HMI tags "DB_SDC_ERROR_STAT_EMS011"
   "DB_SDC_ERRORS_STAT_ER_AKT[11].ER_TRIGER" : Word = PLC DB_SDC_ERRORS_STAT.ER_AKT[11].ER_TRIGER AT %DB3724.DBW28680, 1 s
   "DB_SDC_ERRORS_STAT_ER_AKT[11].ER_STAT[1].DRIVE_POS" : DInt = PLC DB_SDC_ERRORS_STAT.ER_AKT[11].ER_STAT[1].DRIVE_POS AT %DB3724.DBD28686, 1 s
   "DB_SDC_ERRORS_STAT_ER_AKT[11].ER_STAT[1].ERROR" : Int = PLC DB_SDC_ERRORS_STAT.ER_AKT[11].ER_STAT[1].ERROR AT %DB3724.DBW28692, 1 s
   "DB_SDC_ERRORS_STAT_ER_AKT[11].ER_STAT[2].DRIVE_POS" : DInt = PLC DB_SDC_ERRORS_STAT.ER_AKT[11].ER_STAT[2].DRIVE_POS AT %DB3724.DBD28702, 1 s
   "DB_SDC_ERRORS_STAT_ER_AKT[11].ER_STAT[2].ERROR" : Int = PLC DB_SDC_ERRORS_STAT.ER_AKT[59].ER_STAT[4].ERROR AT %DB3724.DBW28708, 1 s
   "DB_SDC_ERRORS_STAT_ER_AKT[11].ER_STAT[3].DRIVE_POS" : DInt = PLC DB_SDC_ERRORS_STAT.ER_AKT[11].ER_STAT[3].DRIVE_POS AT %DB3724.DBD28718, 1 s
   "DB_SDC_ERRORS_STAT_ER_AKT[11].ER_STAT[3].ERROR" : Int = PLC DB_SDC_ERRORS_STAT.ER_AKT[11].ER_STAT[3].ERROR AT %DB3724.DBW28724, 1 s
   "DB_SDC_ERRORS_STAT_ER_AKT[11].ER_STAT[4].DRIVE_POS" : DInt = PLC DB_SDC_ERRORS_STAT.ER_AKT[11].ER_STAT[4].DRIVE_POS AT %DB3724.DBD28734, 1 s
   "DB_SDC_ERRORS_STAT_ER_AKT[11].ER_STAT[4].ERROR" : Int = PLC DB_SDC_ERRORS_STAT.ER_AKT[11].ER_STAT[4].ERROR AT %DB3724.DBW28740, 1 s

HMI tags "DB_SDC_ERROR_STAT_EMS012"
   "DB_SDC_ERRORS_STAT_ER_AKT[12].ER_TRIGER" : Word = PLC DB_SDC_ERRORS_STAT.ER_AKT[12].ER_TRIGER AT %DB3724.DBW28746, 1 s
   "DB_SDC_ERRORS_STAT_ER_AKT[12].ER_STAT[1].DRIVE_POS" : DInt = PLC DB_SDC_ERRORS_STAT.ER_AKT[12].ER_STAT[1].DRIVE_POS AT %DB3724.DBD28752, 1 s
   "DB_SDC_ERRORS_STAT_ER_AKT[12].ER_STAT[1].ERROR" : Int = PLC DB_SDC_ERRORS_STAT.ER_AKT[12].ER_STAT[1].ERROR AT %DB3724.DBW28758, 1 s
   "DB_SDC_ERRORS_STAT_ER_AKT[12].ER_STAT[2].DRIVE_POS" : DInt = PLC DB_SDC_ERRORS_STAT.ER_AKT[12].ER_STAT[2].DRIVE_POS AT %DB3724.DBD28768, 1 s
   "DB_SDC_ERRORS_STAT_ER_AKT[12].ER_STAT[2].ERROR" : Int = PLC DB_SDC_ERRORS_STAT.ER_AKT[12].ER_STAT[2].ERROR AT %DB3724.DBW28774, 1 s
   "DB_SDC_ERRORS_STAT_ER_AKT[12].ER_STAT[3].DRIVE_POS" : DInt = PLC DB_SDC_ERRORS_STAT.ER_AKT[12].ER_STAT[3].DRIVE_POS AT %DB3724.DBD28784, 1 s
   "DB_SDC_ERRORS_STAT_ER_AKT[12].ER_STAT[3].ERROR" : Int = PLC DB_SDC_ERRORS_STAT.ER_AKT[12].ER_STAT[3].ERROR AT %DB3724.DBW28790, 1 s
   "DB_SDC_ERRORS_STAT_ER_AKT[12].ER_STAT[4].DRIVE_POS" : DInt = PLC DB_SDC_ERRORS_STAT.ER_AKT[12].ER_STAT[4].DRIVE_POS AT %DB3724.DBD28800, 1 s
   "DB_SDC_ERRORS_STAT_ER_AKT[12].ER_STAT[4].ERROR" : Int = PLC DB_SDC_ERRORS_STAT.ER_AKT[12].ER_STAT[4].ERROR AT %DB3724.DBW28806, 1 s

HMI tags "DB_SDC_ERROR_STAT_EMS013"
   "DB_SDC_ERRORS_STAT_ER_AKT[13].ER_TRIGER" : Word = PLC DB_SDC_ERRORS_STAT.ER_AKT[13].ER_TRIGER AT %DB3724.DBW28812, 1 s
   "DB_SDC_ERRORS_STAT_ER_AKT[13].ER_STAT[1].DRIVE_POS" : DInt = PLC DB_SDC_ERRORS_STAT.ER_AKT[13].ER_STAT[1].DRIVE_POS AT %DB3724.DBD28818, 1 s
   "DB_SDC_ERRORS_STAT_ER_AKT[13].ER_STAT[1].ERROR" : Int = PLC DB_SDC_ERRORS_STAT.ER_AKT[13].ER_STAT[1].ERROR AT %DB3724.DBW28824, 1 s
   "DB_SDC_ERRORS_STAT_ER_AKT[13].ER_STAT[2].DRIVE_POS" : DInt = PLC DB_SDC_ERRORS_STAT.ER_AKT[13].ER_STAT[2].DRIVE_POS AT %DB3724.DBD28834, 1 s
   "DB_SDC_ERRORS_STAT_ER_AKT[13].ER_STAT[2].ERROR" : Int = PLC DB_SDC_ERRORS_STAT.ER_AKT[13].ER_STAT[2].ERROR AT %DB3724.DBW28840, 1 s
   "DB_SDC_ERRORS_STAT_ER_AKT[13].ER_STAT[3].DRIVE_POS" : DInt = PLC DB_SDC_ERRORS_STAT.ER_AKT[13].ER_STAT[3].DRIVE_POS AT %DB3724.DBD28850, 1 s
   "DB_SDC_ERRORS_STAT_ER_AKT[13].ER_STAT[3].ERROR" : Int = PLC DB_SDC_ERRORS_STAT.ER_AKT[13].ER_STAT[3].ERROR AT %DB3724.DBW28856, 1 s
   "DB_SDC_ERRORS_STAT_ER_AKT[13].ER_STAT[4].DRIVE_POS" : DInt = PLC DB_SDC_ERRORS_STAT.ER_AKT[13].ER_STAT[4].DRIVE_POS AT %DB3724.DBD28866, 1 s
   "DB_SDC_ERRORS_STAT_ER_AKT[13].ER_STAT[4].ERROR" : Int = PLC DB_SDC_ERRORS_STAT.ER_AKT[13].ER_STAT[4].ERROR AT %DB3724.DBW28872, 1 s

HMI tags "DB_SDC_ERROR_STAT_EMS014"
   "DB_SDC_ERRORS_STAT_ER_AKT[14].ER_TRIGER" : Word = PLC DB_SDC_ERRORS_STAT.ER_AKT[14].ER_TRIGER AT %DB3724.DBW28878, 1 s
   "DB_SDC_ERRORS_STAT_ER_AKT[14].ER_STAT[1].DRIVE_POS" : DInt = PLC DB_SDC_ERRORS_STAT.ER_AKT[14].ER_STAT[1].DRIVE_POS AT %DB3724.DBD28884, 1 s
   "DB_SDC_ERRORS_STAT_ER_AKT[14].ER_STAT[1].ERROR" : Int = PLC DB_SDC_ERRORS_STAT.ER_AKT[14].ER_STAT[1].ERROR AT %DB3724.DBW28890, 1 s
   "DB_SDC_ERRORS_STAT_ER_AKT[14].ER_STAT[2].DRIVE_POS" : DInt = PLC DB_SDC_ERRORS_STAT.ER_AKT[14].ER_STAT[2].DRIVE_POS AT %DB3724.DBD28900, 1 s
   "DB_SDC_ERRORS_STAT_ER_AKT[14].ER_STAT[2].ERROR" : Int = PLC DB_SDC_ERRORS_STAT.ER_AKT[14].ER_STAT[2].ERROR AT %DB3724.DBW28906, 1 s
   "DB_SDC_ERRORS_STAT_ER_AKT[14].ER_STAT[3].DRIVE_POS" : DInt = PLC DB_SDC_ERRORS_STAT.ER_AKT[14].ER_STAT[3].DRIVE_POS AT %DB3724.DBD28916, 1 s
   "DB_SDC_ERRORS_STAT_ER_AKT[14].ER_STAT[3].ERROR" : Int = PLC DB_SDC_ERRORS_STAT.ER_AKT[14].ER_STAT[3].ERROR AT %DB3724.DBW28922, 1 s
   "DB_SDC_ERRORS_STAT_ER_AKT[14].ER_STAT[4].DRIVE_POS" : DInt = PLC DB_SDC_ERRORS_STAT.ER_AKT[14].ER_STAT[4].DRIVE_POS AT %DB3724.DBD28932, 1 s
   "DB_SDC_ERRORS_STAT_ER_AKT[14].ER_STAT[4].ERROR" : Int = PLC DB_SDC_ERRORS_STAT.ER_AKT[14].ER_STAT[4].ERROR AT %DB3724.DBW28938, 1 s

HMI tags "DB_SDC_ERROR_STAT_EMS015"
   "DB_SDC_ERRORS_STAT_ER_AKT[15].ER_TRIGER" : Word = PLC DB_SDC_ERRORS_STAT.ER_AKT[15].ER_TRIGER AT %DB3724.DBW28944, 1 s
   "DB_SDC_ERRORS_STAT_ER_AKT[15].ER_STAT[1].DRIVE_POS" : DInt = PLC DB_SDC_ERRORS_STAT.ER_AKT[15].ER_STAT[1].DRIVE_POS AT %DB3724.DBD28950, 1 s
   "DB_SDC_ERRORS_STAT_ER_AKT[15].ER_STAT[1].ERROR" : Int = PLC DB_SDC_ERRORS_STAT.ER_AKT[15].ER_STAT[1].ERROR AT %DB3724.DBW28956, 1 s
   "DB_SDC_ERRORS_STAT_ER_AKT[15].ER_STAT[2].DRIVE_POS" : DInt = PLC DB_SDC_ERRORS_STAT.ER_AKT[15].ER_STAT[2].DRIVE_POS AT %DB3724.DBD28966, 1 s
   "DB_SDC_ERRORS_STAT_ER_AKT[15].ER_STAT[2].ERROR" : Int = PLC DB_SDC_ERRORS_STAT.ER_AKT[15].ER_STAT[2].ERROR AT %DB3724.DBW28972, 1 s
   "DB_SDC_ERRORS_STAT_ER_AKT[15].ER_STAT[3].DRIVE_POS" : DInt = PLC DB_SDC_ERRORS_STAT.ER_AKT[15].ER_STAT[3].DRIVE_POS AT %DB3724.DBD28982, 1 s
   "DB_SDC_ERRORS_STAT_ER_AKT[15].ER_STAT[3].ERROR" : Int = PLC DB_SDC_ERRORS_STAT.ER_AKT[15].ER_STAT[3].ERROR AT %DB3724.DBW28988, 1 s
   "DB_SDC_ERRORS_STAT_ER_AKT[15].ER_STAT[4].DRIVE_POS" : DInt = PLC DB_SDC_ERRORS_STAT.ER_AKT[15].ER_STAT[4].DRIVE_POS AT %DB3724.DBD28998, 1 s
   "DB_SDC_ERRORS_STAT_ER_AKT[15].ER_STAT[4].ERROR" : Int = PLC DB_SDC_ERRORS_STAT.ER_AKT[15].ER_STAT[4].ERROR AT %DB3724.DBW29004, 1 s

HMI tags "DB_SDC_ERROR_STAT_EMS016"
   "DB_SDC_ERRORS_STAT_ER_AKT[16].ER_TRIGER" : Word = PLC DB_SDC_ERRORS_STAT.ER_AKT[16].ER_TRIGER AT %DB3724.DBW29010, 1 s
   "DB_SDC_ERRORS_STAT_ER_AKT[16].ER_STAT[1].DRIVE_POS" : DInt = PLC DB_SDC_ERRORS_STAT.ER_AKT[16].ER_STAT[1].DRIVE_POS AT %DB3724.DBD29016, 1 s
   "DB_SDC_ERRORS_STAT_ER_AKT[16].ER_STAT[1].ERROR" : Int = PLC DB_SDC_ERRORS_STAT.ER_AKT[16].ER_STAT[1].ERROR AT %DB3724.DBW29022, 1 s
   "DB_SDC_ERRORS_STAT_ER_AKT[16].ER_STAT[2].DRIVE_POS" : DInt = PLC DB_SDC_ERRORS_STAT.ER_AKT[16].ER_STAT[2].DRIVE_POS AT %DB3724.DBD29032, 1 s
   "DB_SDC_ERRORS_STAT_ER_AKT[16].ER_STAT[2].ERROR" : Int = PLC DB_SDC_ERRORS_STAT.ER_AKT[16].ER_STAT[2].ERROR AT %DB3724.DBW29038, 1 s
   "DB_SDC_ERRORS_STAT_ER_AKT[16].ER_STAT[3].DRIVE_POS" : DInt = PLC DB_SDC_ERRORS_STAT.ER_AKT[16].ER_STAT[3].DRIVE_POS AT %DB3724.DBD29048, 1 s
   "DB_SDC_ERRORS_STAT_ER_AKT[16].ER_STAT[3].ERROR" : Int = PLC DB_SDC_ERRORS_STAT.ER_AKT[16].ER_STAT[3].ERROR AT %DB3724.DBW29054, 1 s
   "DB_SDC_ERRORS_STAT_ER_AKT[16].ER_STAT[4].DRIVE_POS" : DInt = PLC DB_SDC_ERRORS_STAT.ER_AKT[16].ER_STAT[4].DRIVE_POS AT %DB3724.DBD29064, 1 s
   "DB_SDC_ERRORS_STAT_ER_AKT[16].ER_STAT[4].ERROR" : Int = PLC DB_SDC_ERRORS_STAT.ER_AKT[16].ER_STAT[4].ERROR AT %DB3724.DBW29070, 1 s

HMI tags "DB_SDC_ERROR_STAT_EMS017"
   "DB_SDC_ERRORS_STAT_ER_AKT[17].ER_TRIGER" : Word = PLC DB_SDC_ERRORS_STAT.ER_AKT[17].ER_TRIGER AT %DB3724.DBW29076, 1 s
   "DB_SDC_ERRORS_STAT_ER_AKT[17].ER_STAT[1].DRIVE_POS" : DInt = PLC DB_SDC_ERRORS_STAT.ER_AKT[17].ER_STAT[1].DRIVE_POS AT %DB3724.DBD29082, 1 s
   "DB_SDC_ERRORS_STAT_ER_AKT[17].ER_STAT[1].ERROR" : Int = PLC DB_SDC_ERRORS_STAT.ER_AKT[17].ER_STAT[1].ERROR AT %DB3724.DBW29088, 1 s
   "DB_SDC_ERRORS_STAT_ER_AKT[17].ER_STAT[2].DRIVE_POS" : DInt = PLC DB_SDC_ERRORS_STAT.ER_AKT[17].ER_STAT[2].DRIVE_POS AT %DB3724.DBD29098, 1 s
   "DB_SDC_ERRORS_STAT_ER_AKT[17].ER_STAT[2].ERROR" : Int = PLC DB_SDC_ERRORS_STAT.ER_AKT[17].ER_STAT[2].ERROR AT %DB3724.DBW29104, 1 s
   "DB_SDC_ERRORS_STAT_ER_AKT[17].ER_STAT[3].DRIVE_POS" : DInt = PLC DB_SDC_ERRORS_STAT.ER_AKT[17].ER_STAT[3].DRIVE_POS AT %DB3724.DBD29114, 1 s
   "DB_SDC_ERRORS_STAT_ER_AKT[17].ER_STAT[3].ERROR" : Int = PLC DB_SDC_ERRORS_STAT.ER_AKT[17].ER_STAT[3].ERROR AT %DB3724.DBW29120, 1 s
   "DB_SDC_ERRORS_STAT_ER_AKT[17].ER_STAT[4].DRIVE_POS" : DInt = PLC DB_SDC_ERRORS_STAT.ER_AKT[17].ER_STAT[4].DRIVE_POS AT %DB3724.DBD29130, 1 s
   "DB_SDC_ERRORS_STAT_ER_AKT[17].ER_STAT[4].ERROR" : Int = PLC DB_SDC_ERRORS_STAT.ER_AKT[17].ER_STAT[4].ERROR AT %DB3724.DBW29136, 1 s

HMI tags "DB_SDC_ERROR_STAT_EMS018"
   "DB_SDC_ERRORS_STAT_ER_AKT[18].ER_TRIGER" : Word = PLC DB_SDC_ERRORS_STAT.ER_AKT[18].ER_TRIGER AT %DB3724.DBW29142, 1 s
   "DB_SDC_ERRORS_STAT_ER_AKT[18].ER_STAT[1].DRIVE_POS" : DInt = PLC DB_SDC_ERRORS_STAT.ER_AKT[18].ER_STAT[1].DRIVE_POS AT %DB3724.DBD29148, 1 s
   "DB_SDC_ERRORS_STAT_ER_AKT[18].ER_STAT[1].ERROR" : Int = PLC DB_SDC_ERRORS_STAT.ER_AKT[18].ER_STAT[1].ERROR AT %DB3724.DBW29154, 1 s
   "DB_SDC_ERRORS_STAT_ER_AKT[18].ER_STAT[2].DRIVE_POS" : DInt = PLC DB_SDC_ERRORS_STAT.ER_AKT[18].ER_STAT[2].DRIVE_POS AT %DB3724.DBD29164, 1 s
   "DB_SDC_ERRORS_STAT_ER_AKT[18].ER_STAT[2].ERROR" : Int = PLC DB_SDC_ERRORS_STAT.ER_AKT[18].ER_STAT[2].ERROR AT %DB3724.DBW29170, 1 s
   "DB_SDC_ERRORS_STAT_ER_AKT[18].ER_STAT[3].DRIVE_POS" : DInt = PLC DB_SDC_ERRORS_STAT.ER_AKT[18].ER_STAT[3].DRIVE_POS AT %DB3724.DBD29180, 1 s
   "DB_SDC_ERRORS_STAT_ER_AKT[18].ER_STAT[3].ERROR" : Int = PLC DB_SDC_ERRORS_STAT.ER_AKT[18].ER_STAT[3].ERROR AT %DB3724.DBW29186, 1 s
   "DB_SDC_ERRORS_STAT_ER_AKT[18].ER_STAT[4].DRIVE_POS" : DInt = PLC DB_SDC_ERRORS_STAT.ER_AKT[18].ER_STAT[4].DRIVE_POS AT %DB3724.DBD29196, 1 s
   "DB_SDC_ERRORS_STAT_ER_AKT[18].ER_STAT[4].ERROR" : Int = PLC DB_SDC_ERRORS_STAT.ER_AKT[18].ER_STAT[4].ERROR AT %DB3724.DBW29202, 1 s

HMI tags "DB_SDC_ERROR_STAT_EMS019"
   "DB_SDC_ERRORS_STAT_ER_AKT[19].ER_TRIGER" : Word = PLC DB_SDC_ERRORS_STAT.ER_AKT[19].ER_TRIGER AT %DB3724.DBW29208, 1 s
   "DB_SDC_ERRORS_STAT_ER_AKT[19].ER_STAT[1].DRIVE_POS" : DInt = PLC DB_SDC_ERRORS_STAT.ER_AKT[19].ER_STAT[1].DRIVE_POS AT %DB3724.DBD29214, 1 s
   "DB_SDC_ERRORS_STAT_ER_AKT[19].ER_STAT[1].ERROR" : Int = PLC DB_SDC_ERRORS_STAT.ER_AKT[19].ER_STAT[1].ERROR AT %DB3724.DBW29220, 1 s
   "DB_SDC_ERRORS_STAT_ER_AKT[19].ER_STAT[2].DRIVE_POS" : DInt = PLC DB_SDC_ERRORS_STAT.ER_AKT[19].ER_STAT[2].DRIVE_POS AT %DB3724.DBD29230, 1 s
   "DB_SDC_ERRORS_STAT_ER_AKT[19].ER_STAT[2].ERROR" : Int = PLC DB_SDC_ERRORS_STAT.ER_AKT[19].ER_STAT[2].ERROR AT %DB3724.DBW29236, 1 s
   "DB_SDC_ERRORS_STAT_ER_AKT[19].ER_STAT[3].DRIVE_POS" : DInt = PLC DB_SDC_ERRORS_STAT.ER_AKT[19].ER_STAT[3].DRIVE_POS AT %DB3724.DBD29246, 1 s
   "DB_SDC_ERRORS_STAT_ER_AKT[19].ER_STAT[3].ERROR" : Int = PLC DB_SDC_ERRORS_STAT.ER_AKT[19].ER_STAT[3].ERROR AT %DB3724.DBW29252, 1 s
   "DB_SDC_ERRORS_STAT_ER_AKT[19].ER_STAT[4].DRIVE_POS" : DInt = PLC DB_SDC_ERRORS_STAT.ER_AKT[19].ER_STAT[4].DRIVE_POS AT %DB3724.DBD29262, 1 s
   "DB_SDC_ERRORS_STAT_ER_AKT[19].ER_STAT[4].ERROR" : Int = PLC DB_SDC_ERRORS_STAT.ER_AKT[19].ER_STAT[4].ERROR AT %DB3724.DBW29268, 1 s

HMI tags "DB_SDC_ERROR_STAT_EMS020"
   "DB_SDC_ERRORS_STAT_ER_AKT[20].ER_TRIGER" : Word = PLC DB_SDC_ERRORS_STAT.ER_AKT[20].ER_TRIGER AT %DB3724.DBW29274, 1 s
   "DB_SDC_ERRORS_STAT_ER_AKT[20].ER_STAT[1].DRIVE_POS" : DInt = PLC DB_SDC_ERRORS_STAT.ER_AKT[20].ER_STAT[1].DRIVE_POS AT %DB3724.DBD29280, 1 s
   "DB_SDC_ERRORS_STAT_ER_AKT[20].ER_STAT[1].ERROR" : Int = PLC DB_SDC_ERRORS_STAT.ER_AKT[20].ER_STAT[1].ERROR AT %DB3724.DBW29286, 1 s
   "DB_SDC_ERRORS_STAT_ER_AKT[20].ER_STAT[2].DRIVE_POS" : DInt = PLC DB_SDC_ERRORS_STAT.ER_AKT[20].ER_STAT[2].DRIVE_POS AT %DB3724.DBD29296, 1 s
   "DB_SDC_ERRORS_STAT_ER_AKT[20].ER_STAT[2].ERROR" : Int = PLC DB_SDC_ERRORS_STAT.ER_AKT[20].ER_STAT[2].ERROR AT %DB3724.DBW29302, 1 s
   "DB_SDC_ERRORS_STAT_ER_AKT[20].ER_STAT[3].DRIVE_POS" : DInt = PLC DB_SDC_ERRORS_STAT.ER_AKT[20].ER_STAT[3].DRIVE_POS AT %DB3724.DBD29312, 1 s
   "DB_SDC_ERRORS_STAT_ER_AKT[20].ER_STAT[3].ERROR" : Int = PLC DB_SDC_ERRORS_STAT.ER_AKT[20].ER_STAT[3].ERROR AT %DB3724.DBW29318, 1 s
   "DB_SDC_ERRORS_STAT_ER_AKT[20].ER_STAT[4].DRIVE_POS" : DInt = PLC DB_SDC_ERRORS_STAT.ER_AKT[20].ER_STAT[4].DRIVE_POS AT %DB3724.DBD29328, 1 s
   "DB_SDC_ERRORS_STAT_ER_AKT[20].ER_STAT[4].ERROR" : Int = PLC DB_SDC_ERRORS_STAT.ER_AKT[20].ER_STAT[4].ERROR AT %DB3724.DBW29334, 1 s

HMI tags "DB_SDC_ERROR_STAT_EMS021"
   "DB_SDC_ERRORS_STAT_ER_AKT[21].ER_TRIGER" : Word = PLC DB_SDC_ERRORS_STAT.ER_AKT[21].ER_TRIGER AT %DB3724.DBW29340, 1 s
   "DB_SDC_ERRORS_STAT_ER_AKT[21].ER_STAT[1].DRIVE_POS" : DInt = PLC DB_SDC_ERRORS_STAT.ER_AKT[21].ER_STAT[1].DRIVE_POS AT %DB3724.DBD29346, 1 s
   "DB_SDC_ERRORS_STAT_ER_AKT[21].ER_STAT[1].ERROR" : Int = PLC DB_SDC_ERRORS_STAT.ER_AKT[21].ER_STAT[1].ERROR AT %DB3724.DBW29352, 1 s
   "DB_SDC_ERRORS_STAT_ER_AKT[21].ER_STAT[2].DRIVE_POS" : DInt = PLC DB_SDC_ERRORS_STAT.ER_AKT[21].ER_STAT[2].DRIVE_POS AT %DB3724.DBD29362, 1 s
   "DB_SDC_ERRORS_STAT_ER_AKT[21].ER_STAT[2].ERROR" : Int = PLC DB_SDC_ERRORS_STAT.ER_AKT[21].ER_STAT[2].ERROR AT %DB3724.DBW29368, 1 s
   "DB_SDC_ERRORS_STAT_ER_AKT[21].ER_STAT[3].DRIVE_POS" : DInt = PLC DB_SDC_ERRORS_STAT.ER_AKT[21].ER_STAT[3].DRIVE_POS AT %DB3724.DBD29378, 1 s
   "DB_SDC_ERRORS_STAT_ER_AKT[21].ER_STAT[3].ERROR" : Int = PLC DB_SDC_ERRORS_STAT.ER_AKT[21].ER_STAT[3].ERROR AT %DB3724.DBW29384, 1 s
   "DB_SDC_ERRORS_STAT_ER_AKT[21].ER_STAT[4].DRIVE_POS" : DInt = PLC DB_SDC_ERRORS_STAT.ER_AKT[21].ER_STAT[4].DRIVE_POS AT %DB3724.DBD29394, 1 s
   "DB_SDC_ERRORS_STAT_ER_AKT[21].ER_STAT[4].ERROR" : Int = PLC DB_SDC_ERRORS_STAT.ER_AKT[21].ER_STAT[4].ERROR AT %DB3724.DBW29400, 1 s

HMI tags "DB_SDC_ERROR_STAT_EMS022"
   "DB_SDC_ERRORS_STAT_ER_AKT[22].ER_TRIGER" : Word = PLC DB_SDC_ERRORS_STAT.ER_AKT[22].ER_TRIGER AT %DB3724.DBW29406, 1 s
   "DB_SDC_ERRORS_STAT_ER_AKT[22].ER_STAT[1].DRIVE_POS" : DInt = PLC DB_SDC_ERRORS_STAT.ER_AKT[22].ER_STAT[1].DRIVE_POS AT %DB3724.DBD29412, 1 s
   "DB_SDC_ERRORS_STAT_ER_AKT[22].ER_STAT[1].ERROR" : Int = PLC DB_SDC_ERRORS_STAT.ER_AKT[22].ER_STAT[1].ERROR AT %DB3724.DBW29418, 1 s
   "DB_SDC_ERRORS_STAT_ER_AKT[22].ER_STAT[2].DRIVE_POS" : DInt = PLC DB_SDC_ERRORS_STAT.ER_AKT[22].ER_STAT[2].DRIVE_POS AT %DB3724.DBD29428, 1 s
   "DB_SDC_ERRORS_STAT_ER_AKT[22].ER_STAT[2].ERROR" : Int = PLC DB_SDC_ERRORS_STAT.ER_AKT[22].ER_STAT[2].ERROR AT %DB3724.DBW29434, 1 s
   "DB_SDC_ERRORS_STAT_ER_AKT[22].ER_STAT[3].DRIVE_POS" : DInt = PLC DB_SDC_ERRORS_STAT.ER_AKT[22].ER_STAT[3].DRIVE_POS AT %DB3724.DBD29444, 1 s
   "DB_SDC_ERRORS_STAT_ER_AKT[22].ER_STAT[3].ERROR" : Int = PLC DB_SDC_ERRORS_STAT.ER_AKT[22].ER_STAT[3].ERROR AT %DB3724.DBW29450, 1 s
   "DB_SDC_ERRORS_STAT_ER_AKT[22].ER_STAT[4].DRIVE_POS" : DInt = PLC DB_SDC_ERRORS_STAT.ER_AKT[22].ER_STAT[4].DRIVE_POS AT %DB3724.DBD29460, 1 s
   "DB_SDC_ERRORS_STAT_ER_AKT[22].ER_STAT[4].ERROR" : Int = PLC DB_SDC_ERRORS_STAT.ER_AKT[22].ER_STAT[4].ERROR AT %DB3724.DBW29466, 1 s

HMI tags "DB_SDC_ERROR_STAT_EMS023"
   "DB_SDC_ERRORS_STAT_ER_AKT[23].ER_TRIGER" : Word = PLC DB_SDC_ERRORS_STAT.ER_AKT[23].ER_TRIGER AT %DB3724.DBW29472, 1 s
   "DB_SDC_ERRORS_STAT_ER_AKT[23].ER_STAT[1].DRIVE_POS" : DInt = PLC DB_SDC_ERRORS_STAT.ER_AKT[23].ER_STAT[1].DRIVE_POS AT %DB3724.DBD29478, 1 s
   "DB_SDC_ERRORS_STAT_ER_AKT[23].ER_STAT[1].ERROR" : Int = PLC DB_SDC_ERRORS_STAT.ER_AKT[23].ER_STAT[1].ERROR AT %DB3724.DBW29484, 1 s
   "DB_SDC_ERRORS_STAT_ER_AKT[23].ER_STAT[2].DRIVE_POS" : DInt = PLC DB_SDC_ERRORS_STAT.ER_AKT[23].ER_STAT[2].DRIVE_POS AT %DB3724.DBD29494, 1 s
   "DB_SDC_ERRORS_STAT_ER_AKT[23].ER_STAT[2].ERROR" : Int = PLC DB_SDC_ERRORS_STAT.ER_AKT[23].ER_STAT[2].ERROR AT %DB3724.DBW29500, 1 s
   "DB_SDC_ERRORS_STAT_ER_AKT[23].ER_STAT[3].DRIVE_POS" : DInt = PLC DB_SDC_ERRORS_STAT.ER_AKT[23].ER_STAT[3].DRIVE_POS AT %DB3724.DBD29510, 1 s
   "DB_SDC_ERRORS_STAT_ER_AKT[23].ER_STAT[3].ERROR" : Int = PLC DB_SDC_ERRORS_STAT.ER_AKT[23].ER_STAT[3].ERROR AT %DB3724.DBW29516, 1 s
   "DB_SDC_ERRORS_STAT_ER_AKT[23].ER_STAT[4].DRIVE_POS" : DInt = PLC DB_SDC_ERRORS_STAT.ER_AKT[23].ER_STAT[4].DRIVE_POS AT %DB3724.DBD29526, 1 s
   "DB_SDC_ERRORS_STAT_ER_AKT[23].ER_STAT[4].ERROR" : Int = PLC DB_SDC_ERRORS_STAT.ER_AKT[23].ER_STAT[4].ERROR AT %DB3724.DBW29532, 1 s

HMI tags "DB_SDC_ERROR_STAT_EMS024"
   "DB_SDC_ERRORS_STAT_ER_AKT[24].ER_TRIGER" : Word = PLC DB_SDC_ERRORS_STAT.ER_AKT[24].ER_TRIGER AT %DB3724.DBW29538, 1 s
   "DB_SDC_ERRORS_STAT_ER_AKT[24].ER_STAT[1].DRIVE_POS" : DInt = PLC DB_SDC_ERRORS_STAT.ER_AKT[24].ER_STAT[1].DRIVE_POS AT %DB3724.DBD29544, 1 s
   "DB_SDC_ERRORS_STAT_ER_AKT[24].ER_STAT[1].ERROR" : Int = PLC DB_SDC_ERRORS_STAT.ER_AKT[24].ER_STAT[1].ERROR AT %DB3724.DBW29550, 1 s
   "DB_SDC_ERRORS_STAT_ER_AKT[24].ER_STAT[2].DRIVE_POS" : DInt = PLC DB_SDC_ERRORS_STAT.ER_AKT[24].ER_STAT[2].DRIVE_POS AT %DB3724.DBD29560, 1 s
   "DB_SDC_ERRORS_STAT_ER_AKT[24].ER_STAT[2].ERROR" : Int = PLC DB_SDC_ERRORS_STAT.ER_AKT[24].ER_STAT[2].ERROR AT %DB3724.DBW29566, 1 s
   "DB_SDC_ERRORS_STAT_ER_AKT[24].ER_STAT[3].DRIVE_POS" : DInt = PLC DB_SDC_ERRORS_STAT.ER_AKT[24].ER_STAT[3].DRIVE_POS AT %DB3724.DBD29576, 1 s
   "DB_SDC_ERRORS_STAT_ER_AKT[24].ER_STAT[3].ERROR" : Int = PLC DB_SDC_ERRORS_STAT.ER_AKT[24].ER_STAT[3].ERROR AT %DB3724.DBW29582, 1 s
   "DB_SDC_ERRORS_STAT_ER_AKT[24].ER_STAT[4].DRIVE_POS" : DInt = PLC DB_SDC_ERRORS_STAT.ER_AKT[24].ER_STAT[4].DRIVE_POS AT %DB3724.DBD29592, 1 s
   "DB_SDC_ERRORS_STAT_ER_AKT[24].ER_STAT[4].ERROR" : Int = PLC DB_SDC_ERRORS_STAT.ER_AKT[24].ER_STAT[4].ERROR AT %DB3724.DBW29598, 1 s

HMI tags "DB_SDC_ERROR_STAT_EMS025"
   "DB_SDC_ERRORS_STAT_ER_AKT[25].ER_TRIGER" : Word = PLC DB_SDC_ERRORS_STAT.ER_AKT[25].ER_TRIGER AT %DB3724.DBW29604, 1 s
   "DB_SDC_ERRORS_STAT_ER_AKT[25].ER_STAT[1].DRIVE_POS" : DInt = PLC DB_SDC_ERRORS_STAT.ER_AKT[25].ER_STAT[1].DRIVE_POS AT %DB3724.DBD29610, 1 s
   "DB_SDC_ERRORS_STAT_ER_AKT[25].ER_STAT[1].ERROR" : Int = PLC DB_SDC_ERRORS_STAT.ER_AKT[25].ER_STAT[1].ERROR AT %DB3724.DBW29616, 1 s
   "DB_SDC_ERRORS_STAT_ER_AKT[25].ER_STAT[2].DRIVE_POS" : DInt = PLC DB_SDC_ERRORS_STAT.ER_AKT[25].ER_STAT[2].DRIVE_POS AT %DB3724.DBD29626, 1 s
   "DB_SDC_ERRORS_STAT_ER_AKT[25].ER_STAT[2].ERROR" : Int = PLC DB_SDC_ERRORS_STAT.ER_AKT[25].ER_STAT[2].ERROR AT %DB3724.DBW29632, 1 s
   "DB_SDC_ERRORS_STAT_ER_AKT[25].ER_STAT[3].DRIVE_POS" : DInt = PLC DB_SDC_ERRORS_STAT.ER_AKT[25].ER_STAT[3].DRIVE_POS AT %DB3724.DBD29642, 1 s
   "DB_SDC_ERRORS_STAT_ER_AKT[25].ER_STAT[3].ERROR" : Int = PLC DB_SDC_ERRORS_STAT.ER_AKT[25].ER_STAT[3].ERROR AT %DB3724.DBW29648, 1 s
   "DB_SDC_ERRORS_STAT_ER_AKT[25].ER_STAT[4].DRIVE_POS" : DInt = PLC DB_SDC_ERRORS_STAT.ER_AKT[25].ER_STAT[4].DRIVE_POS AT %DB3724.DBD29658, 1 s
   "DB_SDC_ERRORS_STAT_ER_AKT[25].ER_STAT[4].ERROR" : Int = PLC DB_SDC_ERRORS_STAT.ER_AKT[25].ER_STAT[4].ERROR AT %DB3724.DBW29664, 1 s

HMI tags "DB_SDC_ERROR_STAT_EMS026"
   "DB_SDC_ERRORS_STAT_ER_AKT[26].ER_TRIGER" : Word = PLC DB_SDC_ERRORS_STAT.ER_AKT[26].ER_TRIGER AT %DB3724.DBW29670, 1 s
   "DB_SDC_ERRORS_STAT_ER_AKT[26].ER_STAT[1].DRIVE_POS" : DInt = PLC DB_SDC_ERRORS_STAT.ER_AKT[26].ER_STAT[1].DRIVE_POS AT %DB3724.DBD29676, 1 s
   "DB_SDC_ERRORS_STAT_ER_AKT[26].ER_STAT[1].ERROR" : Int = PLC DB_SDC_ERRORS_STAT.ER_AKT[26].ER_STAT[1].ERROR AT %DB3724.DBW29682, 1 s
   "DB_SDC_ERRORS_STAT_ER_AKT[26].ER_STAT[2].DRIVE_POS" : DInt = PLC DB_SDC_ERRORS_STAT.ER_AKT[26].ER_STAT[2].DRIVE_POS AT %DB3724.DBD29692, 1 s
   "DB_SDC_ERRORS_STAT_ER_AKT[26].ER_STAT[2].ERROR" : Int = PLC DB_SDC_ERRORS_STAT.ER_AKT[26].ER_STAT[2].ERROR AT %DB3724.DBW29698, 1 s
   "DB_SDC_ERRORS_STAT_ER_AKT[26].ER_STAT[3].DRIVE_POS" : DInt = PLC DB_SDC_ERRORS_STAT.ER_AKT[26].ER_STAT[3].DRIVE_POS AT %DB3724.DBD29708, 1 s
   "DB_SDC_ERRORS_STAT_ER_AKT[26].ER_STAT[3].ERROR" : Int = PLC DB_SDC_ERRORS_STAT.ER_AKT[26].ER_STAT[3].ERROR AT %DB3724.DBW29714, 1 s
   "DB_SDC_ERRORS_STAT_ER_AKT[26].ER_STAT[4].DRIVE_POS" : DInt = PLC DB_SDC_ERRORS_STAT.ER_AKT[26].ER_STAT[4].DRIVE_POS AT %DB3724.DBD29724, 1 s
   "DB_SDC_ERRORS_STAT_ER_AKT[26].ER_STAT[4].ERROR" : Int = PLC DB_SDC_ERRORS_STAT.ER_AKT[26].ER_STAT[4].ERROR AT %DB3724.DBW29730, 1 s

HMI tags "DB_SDC_ERROR_STAT_EMS027"
   "DB_SDC_ERRORS_STAT_ER_AKT[27].ER_TRIGER" : Word = PLC DB_SDC_ERRORS_STAT.ER_AKT[27].ER_TRIGER AT %DB3724.DBW29736, 1 s
   "DB_SDC_ERRORS_STAT_ER_AKT[27].ER_STAT[1].DRIVE_POS" : DInt = PLC DB_SDC_ERRORS_STAT.ER_AKT[27].ER_STAT[1].DRIVE_POS AT %DB3724.DBD29742, 1 s
   "DB_SDC_ERRORS_STAT_ER_AKT[27].ER_STAT[1].ERROR" : Int = PLC DB_SDC_ERRORS_STAT.ER_AKT[27].ER_STAT[1].ERROR AT %DB3724.DBW29748, 1 s
   "DB_SDC_ERRORS_STAT_ER_AKT[27].ER_STAT[2].DRIVE_POS" : DInt = PLC DB_SDC_ERRORS_STAT.ER_AKT[27].ER_STAT[2].DRIVE_POS AT %DB3724.DBD29758, 1 s
   "DB_SDC_ERRORS_STAT_ER_AKT[27].ER_STAT[2].ERROR" : Int = PLC DB_SDC_ERRORS_STAT.ER_AKT[27].ER_STAT[2].ERROR AT %DB3724.DBW29764, 1 s
   "DB_SDC_ERRORS_STAT_ER_AKT[27].ER_STAT[3].DRIVE_POS" : DInt = PLC DB_SDC_ERRORS_STAT.ER_AKT[27].ER_STAT[3].DRIVE_POS AT %DB3724.DBD29774, 1 s
   "DB_SDC_ERRORS_STAT_ER_AKT[27].ER_STAT[3].ERROR" : Int = PLC DB_SDC_ERRORS_STAT.ER_AKT[27].ER_STAT[3].ERROR AT %DB3724.DBW29780, 1 s
   "DB_SDC_ERRORS_STAT_ER_AKT[27].ER_STAT[4].DRIVE_POS" : DInt = PLC DB_SDC_ERRORS_STAT.ER_AKT[27].ER_STAT[4].DRIVE_POS AT %DB3724.DBD29790, 1 s
   "DB_SDC_ERRORS_STAT_ER_AKT[27].ER_STAT[4].ERROR" : Int = PLC DB_SDC_ERRORS_STAT.ER_AKT[27].ER_STAT[4].ERROR AT %DB3724.DBW29796, 1 s

HMI tags "DB_SDC_ERROR_STAT_EMS028"
   "DB_SDC_ERRORS_STAT_ER_AKT[28].ER_TRIGER" : Word = PLC DB_SDC_ERRORS_STAT.ER_AKT[28].ER_TRIGER AT %DB3724.DBW29802, 1 s
   "DB_SDC_ERRORS_STAT_ER_AKT[28].ER_STAT[1].DRIVE_POS" : DInt = PLC DB_SDC_ERRORS_STAT.ER_AKT[28].ER_STAT[1].DRIVE_POS AT %DB3724.DBD29808, 1 s
   "DB_SDC_ERRORS_STAT_ER_AKT[28].ER_STAT[1].ERROR" : Int = PLC DB_SDC_ERRORS_STAT.ER_AKT[28].ER_STAT[1].ERROR AT %DB3724.DBW29814, 1 s
   "DB_SDC_ERRORS_STAT_ER_AKT[28].ER_STAT[2].DRIVE_POS" : DInt = PLC DB_SDC_ERRORS_STAT.ER_AKT[28].ER_STAT[2].DRIVE_POS AT %DB3724.DBD29824, 1 s
   "DB_SDC_ERRORS_STAT_ER_AKT[28].ER_STAT[2].ERROR" : Int = PLC DB_SDC_ERRORS_STAT.ER_AKT[28].ER_STAT[2].ERROR AT %DB3724.DBW29830, 1 s
   "DB_SDC_ERRORS_STAT_ER_AKT[28].ER_STAT[3].DRIVE_POS" : DInt = PLC DB_SDC_ERRORS_STAT.ER_AKT[28].ER_STAT[3].DRIVE_POS AT %DB3724.DBD29840, 1 s
   "DB_SDC_ERRORS_STAT_ER_AKT[28].ER_STAT[3].ERROR" : Int = PLC DB_SDC_ERRORS_STAT.ER_AKT[28].ER_STAT[3].ERROR AT %DB3724.DBW29846, 1 s
   "DB_SDC_ERRORS_STAT_ER_AKT[28].ER_STAT[4].DRIVE_POS" : DInt = PLC DB_SDC_ERRORS_STAT.ER_AKT[28].ER_STAT[4].DRIVE_POS AT %DB3724.DBD29856, 1 s
   "DB_SDC_ERRORS_STAT_ER_AKT[28].ER_STAT[4].ERROR" : Int = PLC DB_SDC_ERRORS_STAT.ER_AKT[28].ER_STAT[4].ERROR AT %DB3724.DBW29862, 1 s

HMI tags "DB_SDC_ERROR_STAT_EMS029"
   "DB_SDC_ERRORS_STAT_ER_AKT[29].ER_TRIGER" : Word = PLC DB_SDC_ERRORS_STAT.ER_AKT[29].ER_TRIGER AT %DB3724.DBW29868, 1 s
   "DB_SDC_ERRORS_STAT_ER_AKT[29].ER_STAT[1].DRIVE_POS" : DInt = PLC DB_SDC_ERRORS_STAT.ER_AKT[29].ER_STAT[1].DRIVE_POS AT %DB3724.DBD29874, 1 s
   "DB_SDC_ERRORS_STAT_ER_AKT[29].ER_STAT[1].ERROR" : Int = PLC DB_SDC_ERRORS_STAT.ER_AKT[29].ER_STAT[1].ERROR AT %DB3724.DBW29880, 1 s
   "DB_SDC_ERRORS_STAT_ER_AKT[29].ER_STAT[2].DRIVE_POS" : DInt = PLC DB_SDC_ERRORS_STAT.ER_AKT[29].ER_STAT[2].DRIVE_POS AT %DB3724.DBD29890, 1 s
   "DB_SDC_ERRORS_STAT_ER_AKT[29].ER_STAT[2]" : UDT_SDC_TS_IF_STATUS_VAL = PLC DB_SDC_ERRORS_STAT.ER_AKT[29].ER_STAT[2] AT %DB3724.DBX29886.0, 1 s
   "DB_SDC_ERRORS_STAT_ER_AKT[29].ER_STAT[3].DRIVE_POS" : DInt = PLC DB_SDC_ERRORS_STAT.ER_AKT[29].ER_STAT[3].DRIVE_POS AT %DB3724.DBD29906, 1 s
   "DB_SDC_ERRORS_STAT_ER_AKT[29].ER_STAT[3].ERROR" : Int = PLC DB_SDC_ERRORS_STAT.ER_AKT[29].ER_STAT[3].ERROR AT %DB3724.DBW29912, 1 s
   "DB_SDC_ERRORS_STAT_ER_AKT[29].ER_STAT[4].DRIVE_POS" : DInt = PLC DB_SDC_ERRORS_STAT.ER_AKT[29].ER_STAT[4].DRIVE_POS AT %DB3724.DBD29922, 1 s
   "DB_SDC_ERRORS_STAT_ER_AKT[29].ER_STAT[4].ERROR" : Int = PLC DB_SDC_ERRORS_STAT.ER_AKT[29].ER_STAT[4].ERROR AT %DB3724.DBW29928, 1 s

HMI tags "DB_SDC_ERROR_STAT_EMS030"
   "DB_SDC_ERRORS_STAT_ER_AKT[30].ER_TRIGER" : Word = PLC DB_SDC_ERRORS_STAT.ER_AKT[30].ER_TRIGER AT %DB3724.DBW29934, 1 s
   "DB_SDC_ERRORS_STAT_ER_AKT[30].ER_STAT[1].DRIVE_POS" : DInt = PLC DB_SDC_ERRORS_STAT.ER_AKT[30].ER_STAT[1].DRIVE_POS AT %DB3724.DBD29940, 1 s
   "DB_SDC_ERRORS_STAT_ER_AKT[30].ER_STAT[1].ERROR" : Int = PLC DB_SDC_ERRORS_STAT.ER_AKT[30].ER_STAT[1].ERROR AT %DB3724.DBW29946, 1 s
   "DB_SDC_ERRORS_STAT_ER_AKT[30].ER_STAT[2].DRIVE_POS" : DInt = PLC DB_SDC_ERRORS_STAT.ER_AKT[30].ER_STAT[2].DRIVE_POS AT %DB3724.DBD29956, 1 s
   "DB_SDC_ERRORS_STAT_ER_AKT[30].ER_STAT[2].ERROR" : Int = PLC DB_SDC_ERRORS_STAT.ER_AKT[30].ER_STAT[2].ERROR AT %DB3724.DBW29962, 1 s
   "DB_SDC_ERRORS_STAT_ER_AKT[30].ER_STAT[3].DRIVE_POS" : DInt = PLC DB_SDC_ERRORS_STAT.ER_AKT[30].ER_STAT[3].DRIVE_POS AT %DB3724.DBD29972, 1 s
   "DB_SDC_ERRORS_STAT_ER_AKT[30].ER_STAT[3].ERROR" : Int = PLC DB_SDC_ERRORS_STAT.ER_AKT[30].ER_STAT[3].ERROR AT %DB3724.DBW29978, 1 s
   "DB_SDC_ERRORS_STAT_ER_AKT[30].ER_STAT[4].DRIVE_POS" : DInt = PLC DB_SDC_ERRORS_STAT.ER_AKT[30].ER_STAT[4].DRIVE_POS AT %DB3724.DBD29988, 1 s
   "DB_SDC_ERRORS_STAT_ER_AKT[30].ER_STAT[4].ERROR" : Int = PLC DB_SDC_ERRORS_STAT.ER_AKT[30].ER_STAT[4].ERROR AT %DB3724.DBW29994, 1 s
